VAR_GLOBAL   // PLC tag table "GW_SDC_TO_EMS01_TagTable"
   "SDC_EMS01_Carrier1_Spare0" AT %Q10768.0 : Bool;
   "SDC_EMS01_Carrier1_DriveTripped" AT %Q10768.1 : Bool;
   "SDC_EMS01_Carrier1_Spare2" AT %Q10768.2 : Bool;
   "SDC_EMS01_Carrier1_PositioningComplete" AT %Q10768.3 : Bool;
   "SDC_EMS01_Carrier1_RunStopPressed" AT %Q10768.4 : Bool;
   "SDC_EMS01_Carrier1_Moving" AT %Q10768.5 : Bool;
   "SDC_EMS01_Carrier1_Faulted" AT %Q10768.6 : Bool;
   "SDC_EMS01_Carrier1_InAuto" AT %Q10768.7 : Bool;
   "SDC_EMS01_Carrier2_Spare0" AT %Q10769.0 : Bool;
   "SDC_EMS01_Carrier2_DriveTripped" AT %Q10769.1 : Bool;
   "SDC_EMS01_Carrier2_Spare2" AT %Q10769.2 : Bool;
   "SDC_EMS01_Carrier2_PositioningComplete" AT %Q10769.3 : Bool;
   "SDC_EMS01_Carrier2_RunStopPressed" AT %Q10769.4 : Bool;
   "SDC_EMS01_Carrier2_Moving" AT %Q10769.5 : Bool;
   "SDC_EMS01_Carrier2_Faulted" AT %Q10769.6 : Bool;
   "SDC_EMS01_Carrier2_InAuto" AT %Q10769.7 : Bool;
   "SDC_EMS01_Carrier3_Spare0" AT %Q10770.0 : Bool;
   "SDC_EMS01_Carrier3_DriveTripped" AT %Q10770.1 : Bool;
   "SDC_EMS01_Carrier3_Spare2" AT %Q10770.2 : Bool;
   "SDC_EMS01_Carrier3_PositioningComplete" AT %Q10770.3 : Bool;
   "SDC_EMS01_Carrier3_RunStopPressed" AT %Q10770.4 : Bool;
   "SDC_EMS01_Carrier3_Moving" AT %Q10770.5 : Bool;
   "SDC_EMS01_Carrier3_Faulted" AT %Q10770.6 : Bool;
   "SDC_EMS01_Carrier3_InAuto" AT %Q10770.7 : Bool;
   "SDC_EMS01_Carrier4_Spare0" AT %Q10771.0 : Bool;
   "SDC_EMS01_Carrier4_DriveTripped" AT %Q10771.1 : Bool;
   "SDC_EMS01_Carrier4_Spare2" AT %Q10771.2 : Bool;
   "SDC_EMS01_Carrier4_PositioningComplete" AT %Q10771.3 : Bool;
   "SDC_EMS01_Carrier4_RunStopPressed" AT %Q10771.4 : Bool;
   "SDC_EMS01_Carrier4_Moving" AT %Q10771.5 : Bool;
   "SDC_EMS01_Carrier4_Faulted" AT %Q10771.6 : Bool;
   "SDC_EMS01_Carrier4_InAuto" AT %Q10771.7 : Bool;
   "SDC_EMS01_Carrier5_Spare0" AT %Q10772.0 : Bool;
   "SDC_EMS01_Carrier5_DriveTripped" AT %Q10772.1 : Bool;
   "SDC_EMS01_Carrier5_Spare2" AT %Q10772.2 : Bool;
   "SDC_EMS01_Carrier5_PositioningComplete" AT %Q10772.3 : Bool;
   "SDC_EMS01_Carrier5_RunStopPressed" AT %Q10772.4 : Bool;
   "SDC_EMS01_Carrier5_Moving" AT %Q10772.5 : Bool;
   "SDC_EMS01_Carrier5_Faulted" AT %Q10772.6 : Bool;
   "SDC_EMS01_Carrier5_InAuto" AT %Q10772.7 : Bool;
   "SDC_EMS01_Carrier6_Spare0" AT %Q10773.0 : Bool;
   "SDC_EMS01_Carrier6_DriveTripped" AT %Q10773.1 : Bool;
   "SDC_EMS01_Carrier6_Spare2" AT %Q10773.2 : Bool;
   "SDC_EMS01_Carrier6_PositioningComplete" AT %Q10773.3 : Bool;
   "SDC_EMS01_Carrier6_RunStopPressed" AT %Q10773.4 : Bool;
   "SDC_EMS01_Carrier6_Moving" AT %Q10773.5 : Bool;
   "SDC_EMS01_Carrier6_Faulted" AT %Q10773.6 : Bool;
   "SDC_EMS01_Carrier6_InAuto" AT %Q10773.7 : Bool;
   "SDC_EMS01_Carrier7_Spare0" AT %Q10774.0 : Bool;
   "SDC_EMS01_Carrier7_DriveTripped" AT %Q10774.1 : Bool;
   "SDC_EMS01_Carrier7_Spare2" AT %Q10774.2 : Bool;
   "SDC_EMS01_Carrier7_PositioningComplete" AT %Q10774.3 : Bool;
   "SDC_EMS01_Carrier7_RunStopPressed" AT %Q10774.4 : Bool;
   "SDC_EMS01_Carrier7_Moving" AT %Q10774.5 : Bool;
   "SDC_EMS01_Carrier7_Faulted" AT %Q10774.6 : Bool;
   "SDC_EMS01_Carrier7_InAuto" AT %Q10774.7 : Bool;
   "SDC_EMS01_Carrier8_Spare0" AT %Q10775.0 : Bool;
   "SDC_EMS01_Carrier8_DriveTripped" AT %Q10775.1 : Bool;
   "SDC_EMS01_Carrier8_Spare2" AT %Q10775.2 : Bool;
   "SDC_EMS01_Carrier8_PositioningComplete" AT %Q10775.3 : Bool;
   "SDC_EMS01_Carrier8_RunStopPressed" AT %Q10775.4 : Bool;
   "SDC_EMS01_Carrier8_Moving" AT %Q10775.5 : Bool;
   "SDC_EMS01_Carrier8_Faulted" AT %Q10775.6 : Bool;
   "SDC_EMS01_Carrier8_InAuto" AT %Q10775.7 : Bool;
   "SDC_EMS01_Carrier9_Spare0" AT %Q10776.0 : Bool;
   "SDC_EMS01_Carrier9_DriveTripped" AT %Q10776.1 : Bool;
   "SDC_EMS01_Carrier9_Spare2" AT %Q10776.2 : Bool;
   "SDC_EMS01_Carrier9_PositioningComplete" AT %Q10776.3 : Bool;
   "SDC_EMS01_Carrier9_RunStopPressed" AT %Q10776.4 : Bool;
   "SDC_EMS01_Carrier9_Moving" AT %Q10776.5 : Bool;
   "SDC_EMS01_Carrier9_Faulted" AT %Q10776.6 : Bool;
   "SDC_EMS01_Carrier9_InAuto" AT %Q10776.7 : Bool;
   "SDC_EMS01_Carrier10_Spare0" AT %Q10777.0 : Bool;
   "SDC_EMS01_Carrier10_DriveTripped" AT %Q10777.1 : Bool;
   "SDC_EMS01_Carrier10_Spare2" AT %Q10777.2 : Bool;
   "SDC_EMS01_Carrier10_PositioningComplete" AT %Q10777.3 : Bool;
   "SDC_EMS01_Carrier10_RunStopPressed" AT %Q10777.4 : Bool;
   "SDC_EMS01_Carrier10_Moving" AT %Q10777.5 : Bool;
   "SDC_EMS01_Carrier10_Faulted" AT %Q10777.6 : Bool;
   "SDC_EMS01_Carrier10_InAuto" AT %Q10777.7 : Bool;
   "SDC_EMS01_Carrier11_Spare0" AT %Q10778.0 : Bool;
   "SDC_EMS01_Carrier11_DriveTripped" AT %Q10778.1 : Bool;
   "SDC_EMS01_Carrier11_Spare2" AT %Q10778.2 : Bool;
   "SDC_EMS01_Carrier11_PositioningComplete" AT %Q10778.3 : Bool;
   "SDC_EMS01_Carrier11_RunStopPressed" AT %Q10778.4 : Bool;
   "SDC_EMS01_Carrier11_Moving" AT %Q10778.5 : Bool;
   "SDC_EMS01_Carrier11_Faulted" AT %Q10778.6 : Bool;
   "SDC_EMS01_Carrier11_InAuto" AT %Q10778.7 : Bool;
   "SDC_EMS01_Carrier12_Spare0" AT %Q10779.0 : Bool;
   "SDC_EMS01_Carrier12_DriveTripped" AT %Q10779.1 : Bool;
   "SDC_EMS01_Carrier12_Spare2" AT %Q10779.2 : Bool;
   "SDC_EMS01_Carrier12_PositioningComplete" AT %Q10779.3 : Bool;
   "SDC_EMS01_Carrier12_RunStopPressed" AT %Q10779.4 : Bool;
   "SDC_EMS01_Carrier12_Moving" AT %Q10779.5 : Bool;
   "SDC_EMS01_Carrier12_Faulted" AT %Q10779.6 : Bool;
   "SDC_EMS01_Carrier12_InAuto" AT %Q10779.7 : Bool;
   "SDC_EMS01_Carrier13_Spare0" AT %Q10780.0 : Bool;
   "SDC_EMS01_Carrier13_DriveTripped" AT %Q10780.1 : Bool;
   "SDC_EMS01_Carrier13_Spare2" AT %Q10780.2 : Bool;
   "SDC_EMS01_Carrier13_PositioningComplete" AT %Q10780.3 : Bool;
   "SDC_EMS01_Carrier13_RunStopPressed" AT %Q10780.4 : Bool;
   "SDC_EMS01_Carrier13_Moving" AT %Q10780.5 : Bool;
   "SDC_EMS01_Carrier13_Faulted" AT %Q10780.6 : Bool;
   "SDC_EMS01_Carrier13_InAuto" AT %Q10780.7 : Bool;
   "SDC_EMS01_Carrier14_Spare0" AT %Q10781.0 : Bool;
   "SDC_EMS01_Carrier14_DriveTripped" AT %Q10781.1 : Bool;
   "SDC_EMS01_Carrier14_Spare2" AT %Q10781.2 : Bool;
   "SDC_EMS01_Carrier14_PositioningComplete" AT %Q10781.3 : Bool;
   "SDC_EMS01_Carrier14_RunStopPressed" AT %Q10781.4 : Bool;
   "SDC_EMS01_Carrier14_Moving" AT %Q10781.5 : Bool;
   "SDC_EMS01_Carrier14_Faulted" AT %Q10781.6 : Bool;
   "SDC_EMS01_Carrier14_InAuto" AT %Q10781.7 : Bool;
   "SDC_EMS01_Carrier15_Spare0" AT %Q10782.0 : Bool;
   "SDC_EMS01_Carrier15_DriveTripped" AT %Q10782.1 : Bool;
   "SDC_EMS01_Carrier15_Spare2" AT %Q10782.2 : Bool;
   "SDC_EMS01_Carrier15_PositioningComplete" AT %Q10782.3 : Bool;
   "SDC_EMS01_Carrier15_RunStopPressed" AT %Q10782.4 : Bool;
   "SDC_EMS01_Carrier15_Moving" AT %Q10782.5 : Bool;
   "SDC_EMS01_Carrier15_Faulted" AT %Q10782.6 : Bool;
   "SDC_EMS01_Carrier15_InAuto" AT %Q10782.7 : Bool;
   "SDC_EMS01_Carrier16_Spare0" AT %Q10783.0 : Bool;
   "SDC_EMS01_Carrier16_DriveTripped" AT %Q10783.1 : Bool;
   "SDC_EMS01_Carrier16_Spare2" AT %Q10783.2 : Bool;
   "SDC_EMS01_Carrier16_PositioningComplete" AT %Q10783.3 : Bool;
   "SDC_EMS01_Carrier16_RunStopPressed" AT %Q10783.4 : Bool;
   "SDC_EMS01_Carrier16_Moving" AT %Q10783.5 : Bool;
   "SDC_EMS01_Carrier16_Faulted" AT %Q10783.6 : Bool;
   "SDC_EMS01_Carrier16_InAuto" AT %Q10783.7 : Bool;
   "SDC_EMS01_Carrier17_Spare0" AT %Q10784.0 : Bool;
   "SDC_EMS01_Carrier17_DriveTripped" AT %Q10784.1 : Bool;
   "SDC_EMS01_Carrier17_Spare2" AT %Q10784.2 : Bool;
   "SDC_EMS01_Carrier17_PositioningComplete" AT %Q10784.3 : Bool;
   "SDC_EMS01_Carrier17_RunStopPressed" AT %Q10784.4 : Bool;
   "SDC_EMS01_Carrier17_Moving" AT %Q10784.5 : Bool;
   "SDC_EMS01_Carrier17_Faulted" AT %Q10784.6 : Bool;
   "SDC_EMS01_Carrier17_InAuto" AT %Q10784.7 : Bool;
   "SDC_EMS01_Carrier18_Spare0" AT %Q10785.0 : Bool;
   "SDC_EMS01_Carrier18_DriveTripped" AT %Q10785.1 : Bool;
   "SDC_EMS01_Carrier18_Spare2" AT %Q10785.2 : Bool;
   "SDC_EMS01_Carrier18_PositioningComplete" AT %Q10785.3 : Bool;
   "SDC_EMS01_Carrier18_RunStopPressed" AT %Q10785.4 : Bool;
   "SDC_EMS01_Carrier18_Moving" AT %Q10785.5 : Bool;
   "SDC_EMS01_Carrier18_Faulted" AT %Q10785.6 : Bool;
   "SDC_EMS01_Carrier18_InAuto" AT %Q10785.7 : Bool;
   "SDC_EMS01_Carrier19_Spare0" AT %Q10786.0 : Bool;
   "SDC_EMS01_Carrier19_DriveTripped" AT %Q10786.1 : Bool;
   "SDC_EMS01_Carrier19_Spare2" AT %Q10786.2 : Bool;
   "SDC_EMS01_Carrier19_PositioningComplete" AT %Q10786.3 : Bool;
   "SDC_EMS01_Carrier19_RunStopPressed" AT %Q10786.4 : Bool;
   "SDC_EMS01_Carrier19_Moving" AT %Q10786.5 : Bool;
   "SDC_EMS01_Carrier19_Faulted" AT %Q10786.6 : Bool;
   "SDC_EMS01_Carrier19_InAuto" AT %Q10786.7 : Bool;
   "SDC_EMS01_Carrier20_Spare0" AT %Q10787.0 : Bool;
   "SDC_EMS01_Carrier20_DriveTripped" AT %Q10787.1 : Bool;
   "SDC_EMS01_Carrier20_Spare2" AT %Q10787.2 : Bool;
   "SDC_EMS01_Carrier20_PositioningComplete" AT %Q10787.3 : Bool;
   "SDC_EMS01_Carrier20_RunStopPressed" AT %Q10787.4 : Bool;
   "SDC_EMS01_Carrier20_Moving" AT %Q10787.5 : Bool;
   "SDC_EMS01_Carrier20_Faulted" AT %Q10787.6 : Bool;
   "SDC_EMS01_Carrier20_InAuto" AT %Q10787.7 : Bool;
   "SDC_EMS01_Carrier21_Spare0" AT %Q10788.0 : Bool;
   "SDC_EMS01_Carrier21_DriveTripped" AT %Q10788.1 : Bool;
   "SDC_EMS01_Carrier21_Spare2" AT %Q10788.2 : Bool;
   "SDC_EMS01_Carrier21_PositioningComplete" AT %Q10788.3 : Bool;
   "SDC_EMS01_Carrier21_RunStopPressed" AT %Q10788.4 : Bool;
   "SDC_EMS01_Carrier21_Moving" AT %Q10788.5 : Bool;
   "SDC_EMS01_Carrier21_Faulted" AT %Q10788.6 : Bool;
   "SDC_EMS01_Carrier21_InAuto" AT %Q10788.7 : Bool;
   "SDC_EMS01_Carrier22_Spare0" AT %Q10789.0 : Bool;
   "SDC_EMS01_Carrier22_DriveTripped" AT %Q10789.1 : Bool;
   "SDC_EMS01_Carrier22_Spare2" AT %Q10789.2 : Bool;
   "SDC_EMS01_Carrier22_PositioningComplete" AT %Q10789.3 : Bool;
   "SDC_EMS01_Carrier22_RunStopPressed" AT %Q10789.4 : Bool;
   "SDC_EMS01_Carrier22_Moving" AT %Q10789.5 : Bool;
   "SDC_EMS01_Carrier22_Faulted" AT %Q10789.6 : Bool;
   "SDC_EMS01_Carrier22_InAuto" AT %Q10789.7 : Bool;
   "SDC_EMS01_Carrier23_Spare0" AT %Q10790.0 : Bool;
   "SDC_EMS01_Carrier23_DriveTripped" AT %Q10790.1 : Bool;
   "SDC_EMS01_Carrier23_Spare2" AT %Q10790.2 : Bool;
   "SDC_EMS01_Carrier23_PositioningComplete" AT %Q10790.3 : Bool;
   "SDC_EMS01_Carrier23_RunStopPressed" AT %Q10790.4 : Bool;
   "SDC_EMS01_Carrier23_Moving" AT %Q10790.5 : Bool;
   "SDC_EMS01_Carrier23_Faulted" AT %Q10790.6 : Bool;
   "SDC_EMS01_Carrier23_InAuto" AT %Q10790.7 : Bool;
   "SDC_EMS01_Carrier24_Spare0" AT %Q10791.0 : Bool;
   "SDC_EMS01_Carrier24_DriveTripped" AT %Q10791.1 : Bool;
   "SDC_EMS01_Carrier24_Spare2" AT %Q10791.2 : Bool;
   "SDC_EMS01_Carrier24_PositioningComplete" AT %Q10791.3 : Bool;
   "SDC_EMS01_Carrier24_RunStopPressed" AT %Q10791.4 : Bool;
   "SDC_EMS01_Carrier24_Moving" AT %Q10791.5 : Bool;
   "SDC_EMS01_Carrier24_Faulted" AT %Q10791.6 : Bool;
   "SDC_EMS01_Carrier24_InAuto" AT %Q10791.7 : Bool;
   "SDC_EMS01_Carrier25_Spare0" AT %Q10792.0 : Bool;
   "SDC_EMS01_Carrier25_DriveTripped" AT %Q10792.1 : Bool;
   "SDC_EMS01_Carrier25_Spare2" AT %Q10792.2 : Bool;
   "SDC_EMS01_Carrier25_PositioningComplete" AT %Q10792.3 : Bool;
   "SDC_EMS01_Carrier25_RunStopPressed" AT %Q10792.4 : Bool;
   "SDC_EMS01_Carrier25_Moving" AT %Q10792.5 : Bool;
   "SDC_EMS01_Carrier25_Faulted" AT %Q10792.6 : Bool;
   "SDC_EMS01_Carrier25_InAuto" AT %Q10792.7 : Bool;
   "SDC_EMS01_Carrier26_Spare0" AT %Q10793.0 : Bool;
   "SDC_EMS01_Carrier26_DriveTripped" AT %Q10793.1 : Bool;
   "SDC_EMS01_Carrier26_Spare2" AT %Q10793.2 : Bool;
   "SDC_EMS01_Carrier26_PositioningComplete" AT %Q10793.3 : Bool;
   "SDC_EMS01_Carrier26_RunStopPressed" AT %Q10793.4 : Bool;
   "SDC_EMS01_Carrier26_Moving" AT %Q10793.5 : Bool;
   "SDC_EMS01_Carrier26_Faulted" AT %Q10793.6 : Bool;
   "SDC_EMS01_Carrier26_InAuto" AT %Q10793.7 : Bool;
   "SDC_EMS01_Carrier27_Spare0" AT %Q10794.0 : Bool;
   "SDC_EMS01_Carrier27_DriveTripped" AT %Q10794.1 : Bool;
   "SDC_EMS01_Carrier27_Spare2" AT %Q10794.2 : Bool;
   "SDC_EMS01_Carrier27_PositioningComplete" AT %Q10794.3 : Bool;
   "SDC_EMS01_Carrier27_RunStopPressed" AT %Q10794.4 : Bool;
   "SDC_EMS01_Carrier27_Moving" AT %Q10794.5 : Bool;
   "SDC_EMS01_Carrier27_Faulted" AT %Q10794.6 : Bool;
   "SDC_EMS01_Carrier27_InAuto" AT %Q10794.7 : Bool;
   "SDC_EMS01_Carrier28_Spare0" AT %Q10795.0 : Bool;
   "SDC_EMS01_Carrier28_DriveTripped" AT %Q10795.1 : Bool;
   "SDC_EMS01_Carrier28_Spare2" AT %Q10795.2 : Bool;
   "SDC_EMS01_Carrier28_PositioningComplete" AT %Q10795.3 : Bool;
   "SDC_EMS01_Carrier28_RunStopPressed" AT %Q10795.4 : Bool;
   "SDC_EMS01_Carrier28_Moving" AT %Q10795.5 : Bool;
   "SDC_EMS01_Carrier28_Faulted" AT %Q10795.6 : Bool;
   "SDC_EMS01_Carrier28_InAuto" AT %Q10795.7 : Bool;
   "SDC_EMS01_Carrier29_Spare0" AT %Q10796.0 : Bool;
   "SDC_EMS01_Carrier29_DriveTripped" AT %Q10796.1 : Bool;
   "SDC_EMS01_Carrier29_Spare2" AT %Q10796.2 : Bool;
   "SDC_EMS01_Carrier29_PositioningComplete" AT %Q10796.3 : Bool;
   "SDC_EMS01_Carrier29_RunStopPressed" AT %Q10796.4 : Bool;
   "SDC_EMS01_Carrier29_Moving" AT %Q10796.5 : Bool;
   "SDC_EMS01_Carrier29_Faulted" AT %Q10796.6 : Bool;
   "SDC_EMS01_Carrier29_InAuto" AT %Q10796.7 : Bool;
   "SDC_EMS01_Carrier30_Spare0" AT %Q10797.0 : Bool;
   "SDC_EMS01_Carrier30_DriveTripped" AT %Q10797.1 : Bool;
   "SDC_EMS01_Carrier30_Spare2" AT %Q10797.2 : Bool;
   "SDC_EMS01_Carrier30_PositioningComplete" AT %Q10797.3 : Bool;
   "SDC_EMS01_Carrier30_RunStopPressed" AT %Q10797.4 : Bool;
   "SDC_EMS01_Carrier30_Moving" AT %Q10797.5 : Bool;
   "SDC_EMS01_Carrier30_Faulted" AT %Q10797.6 : Bool;
   "SDC_EMS01_Carrier30_InAuto" AT %Q10797.7 : Bool;
   "SDC_EMS01_Carrier31_Spare0" AT %Q10798.0 : Bool;
   "SDC_EMS01_Carrier31_DriveTripped" AT %Q10798.1 : Bool;
   "SDC_EMS01_Carrier31_Spare2" AT %Q10798.2 : Bool;
   "SDC_EMS01_Carrier31_PositioningComplete" AT %Q10798.3 : Bool;
   "SDC_EMS01_Carrier31_RunStopPressed" AT %Q10798.4 : Bool;
   "SDC_EMS01_Carrier31_Moving" AT %Q10798.5 : Bool;
   "SDC_EMS01_Carrier31_Faulted" AT %Q10798.6 : Bool;
   "SDC_EMS01_Carrier31_InAuto" AT %Q10798.7 : Bool;
   "SDC_EMS01_Carrier32_Spare0" AT %Q10799.0 : Bool;
   "SDC_EMS01_Carrier32_DriveTripped" AT %Q10799.1 : Bool;
   "SDC_EMS01_Carrier32_Spare2" AT %Q10799.2 : Bool;
   "SDC_EMS01_Carrier32_PositioningComplete" AT %Q10799.3 : Bool;
   "SDC_EMS01_Carrier32_RunStopPressed" AT %Q10799.4 : Bool;
   "SDC_EMS01_Carrier32_Moving" AT %Q10799.5 : Bool;
   "SDC_EMS01_Carrier32_Faulted" AT %Q10799.6 : Bool;
   "SDC_EMS01_Carrier32_InAuto" AT %Q10799.7 : Bool;
   "SDC_EMS01_Carrier33_Spare0" AT %Q10800.0 : Bool;
   "SDC_EMS01_Carrier33_DriveTripped" AT %Q10800.1 : Bool;
   "SDC_EMS01_Carrier33_Spare2" AT %Q10800.2 : Bool;
   "SDC_EMS01_Carrier33_PositioningComplete" AT %Q10800.3 : Bool;
   "SDC_EMS01_Carrier33_RunStopPressed" AT %Q10800.4 : Bool;
   "SDC_EMS01_Carrier33_Moving" AT %Q10800.5 : Bool;
   "SDC_EMS01_Carrier33_Faulted" AT %Q10800.6 : Bool;
   "SDC_EMS01_Carrier33_InAuto" AT %Q10800.7 : Bool;
   "SDC_EMS01_Carrier34_Spare0" AT %Q10801.0 : Bool;
   "SDC_EMS01_Carrier34_DriveTripped" AT %Q10801.1 : Bool;
   "SDC_EMS01_Carrier34_Spare2" AT %Q10801.2 : Bool;
   "SDC_EMS01_Carrier34_PositioningComplete" AT %Q10801.3 : Bool;
   "SDC_EMS01_Carrier34_RunStopPressed" AT %Q10801.4 : Bool;
   "SDC_EMS01_Carrier34_Moving" AT %Q10801.5 : Bool;
   "SDC_EMS01_Carrier34_Faulted" AT %Q10801.6 : Bool;
   "SDC_EMS01_Carrier34_InAuto" AT %Q10801.7 : Bool;
   "SDC_EMS01_Carrier35_Spare0" AT %Q10802.0 : Bool;
   "SDC_EMS01_Carrier35_DriveTripped" AT %Q10802.1 : Bool;
   "SDC_EMS01_Carrier35_Spare2" AT %Q10802.2 : Bool;
   "SDC_EMS01_Carrier35_PositioningComplete" AT %Q10802.3 : Bool;
   "SDC_EMS01_Carrier35_RunStopPressed" AT %Q10802.4 : Bool;
   "SDC_EMS01_Carrier35_Moving" AT %Q10802.5 : Bool;
   "SDC_EMS01_Carrier35_Faulted" AT %Q10802.6 : Bool;
   "SDC_EMS01_Carrier35_InAuto" AT %Q10802.7 : Bool;
   "SDC_EMS01_Carrier36_Spare0" AT %Q10803.0 : Bool;
   "SDC_EMS01_Carrier36_DriveTripped" AT %Q10803.1 : Bool;
   "SDC_EMS01_Carrier36_Spare2" AT %Q10803.2 : Bool;
   "SDC_EMS01_Carrier36_PositioningComplete" AT %Q10803.3 : Bool;
   "SDC_EMS01_Carrier36_RunStopPressed" AT %Q10803.4 : Bool;
   "SDC_EMS01_Carrier36_Moving" AT %Q10803.5 : Bool;
   "SDC_EMS01_Carrier36_Faulted" AT %Q10803.6 : Bool;
   "SDC_EMS01_Carrier36_InAuto" AT %Q10803.7 : Bool;
   "SDC_EMS01_Carrier37_Spare0" AT %Q10804.0 : Bool;
   "SDC_EMS01_Carrier37_DriveTripped" AT %Q10804.1 : Bool;
   "SDC_EMS01_Carrier37_Spare2" AT %Q10804.2 : Bool;
   "SDC_EMS01_Carrier37_PositioningComplete" AT %Q10804.3 : Bool;
   "SDC_EMS01_Carrier37_RunStopPressed" AT %Q10804.4 : Bool;
   "SDC_EMS01_Carrier37_Moving" AT %Q10804.5 : Bool;
   "SDC_EMS01_Carrier37_Faulted" AT %Q10804.6 : Bool;
   "SDC_EMS01_Carrier37_InAuto" AT %Q10804.7 : Bool;
   "SDC_EMS01_Carrier38_Spare0" AT %Q10805.0 : Bool;
   "SDC_EMS01_Carrier38_DriveTripped" AT %Q10805.1 : Bool;
   "SDC_EMS01_Carrier38_Spare2" AT %Q10805.2 : Bool;
   "SDC_EMS01_Carrier38_PositioningComplete" AT %Q10805.3 : Bool;
   "SDC_EMS01_Carrier38_RunStopPressed" AT %Q10805.4 : Bool;
   "SDC_EMS01_Carrier38_Moving" AT %Q10805.5 : Bool;
   "SDC_EMS01_Carrier38_Faulted" AT %Q10805.6 : Bool;
   "SDC_EMS01_Carrier38_InAuto" AT %Q10805.7 : Bool;
   "SDC_EMS01_Carrier39_Spare0" AT %Q10806.0 : Bool;
   "SDC_EMS01_Carrier39_DriveTripped" AT %Q10806.1 : Bool;
   "SDC_EMS01_Carrier39_Spare2" AT %Q10806.2 : Bool;
   "SDC_EMS01_Carrier39_PositioningComplete" AT %Q10806.3 : Bool;
   "SDC_EMS01_Carrier39_RunStopPressed" AT %Q10806.4 : Bool;
   "SDC_EMS01_Carrier39_Moving" AT %Q10806.5 : Bool;
   "SDC_EMS01_Carrier39_Faulted" AT %Q10806.6 : Bool;
   "SDC_EMS01_Carrier39_InAuto" AT %Q10806.7 : Bool;
   "SDC_EMS01_Carrier40_Spare0" AT %Q10807.0 : Bool;
   "SDC_EMS01_Carrier40_DriveTripped" AT %Q10807.1 : Bool;
   "SDC_EMS01_Carrier40_Spare2" AT %Q10807.2 : Bool;
   "SDC_EMS01_Carrier40_PositioningComplete" AT %Q10807.3 : Bool;
   "SDC_EMS01_Carrier40_RunStopPressed" AT %Q10807.4 : Bool;
   "SDC_EMS01_Carrier40_Moving" AT %Q10807.5 : Bool;
   "SDC_EMS01_Carrier40_Faulted" AT %Q10807.6 : Bool;
   "SDC_EMS01_Carrier40_InAuto" AT %Q10807.7 : Bool;
   "SDC_EMS01_Carrier41_Spare0" AT %Q10808.0 : Bool;
   "SDC_EMS01_Carrier41_DriveTripped" AT %Q10808.1 : Bool;
   "SDC_EMS01_Carrier41_Spare2" AT %Q10808.2 : Bool;
   "SDC_EMS01_Carrier41_PositioningComplete" AT %Q10808.3 : Bool;
   "SDC_EMS01_Carrier41_RunStopPressed" AT %Q10808.4 : Bool;
   "SDC_EMS01_Carrier41_Moving" AT %Q10808.5 : Bool;
   "SDC_EMS01_Carrier41_Faulted" AT %Q10808.6 : Bool;
   "SDC_EMS01_Carrier41_InAuto" AT %Q10808.7 : Bool;
   "SDC_EMS01_Carrier42_Spare0" AT %Q10809.0 : Bool;
   "SDC_EMS01_Carrier42_DriveTripped" AT %Q10809.1 : Bool;
   "SDC_EMS01_Carrier42_Spare2" AT %Q10809.2 : Bool;
   "SDC_EMS01_Carrier42_PositioningComplete" AT %Q10809.3 : Bool;
   "SDC_EMS01_Carrier42_RunStopPressed" AT %Q10809.4 : Bool;
   "SDC_EMS01_Carrier42_Moving" AT %Q10809.5 : Bool;
   "SDC_EMS01_Carrier42_Faulted" AT %Q10809.6 : Bool;
   "SDC_EMS01_Carrier42_InAuto" AT %Q10809.7 : Bool;
   "SDC_EMS01_Carrier43_Spare0" AT %Q10810.0 : Bool;
   "SDC_EMS01_Carrier43_DriveTripped" AT %Q10810.1 : Bool;
   "SDC_EMS01_Carrier43_Spare2" AT %Q10810.2 : Bool;
   "SDC_EMS01_Carrier43_PositioningComplete" AT %Q10810.3 : Bool;
   "SDC_EMS01_Carrier43_RunStopPressed" AT %Q10810.4 : Bool;
   "SDC_EMS01_Carrier43_Moving" AT %Q10810.5 : Bool;
   "SDC_EMS01_Carrier43_Faulted" AT %Q10810.6 : Bool;
   "SDC_EMS01_Carrier43_InAuto" AT %Q10810.7 : Bool;
   "SDC_EMS01_Carrier44_Spare0" AT %Q10811.0 : Bool;
   "SDC_EMS01_Carrier44_DriveTripped" AT %Q10811.1 : Bool;
   "SDC_EMS01_Carrier44_Spare2" AT %Q10811.2 : Bool;
   "SDC_EMS01_Carrier44_PositioningComplete" AT %Q10811.3 : Bool;
   "SDC_EMS01_Carrier44_RunStopPressed" AT %Q10811.4 : Bool;
   "SDC_EMS01_Carrier44_Moving" AT %Q10811.5 : Bool;
   "SDC_EMS01_Carrier44_Faulted" AT %Q10811.6 : Bool;
   "SDC_EMS01_Carrier44_InAuto" AT %Q10811.7 : Bool;
   "SDC_EMS01_Carrier45_Spare0" AT %Q10812.0 : Bool;
   "SDC_EMS01_Carrier45_DriveTripped" AT %Q10812.1 : Bool;
   "SDC_EMS01_Carrier45_Spare2" AT %Q10812.2 : Bool;
   "SDC_EMS01_Carrier45_PositioningComplete" AT %Q10812.3 : Bool;
   "SDC_EMS01_Carrier45_RunStopPressed" AT %Q10812.4 : Bool;
   "SDC_EMS01_Carrier45_Moving" AT %Q10812.5 : Bool;
   "SDC_EMS01_Carrier45_Faulted" AT %Q10812.6 : Bool;
   "SDC_EMS01_Carrier45_InAuto" AT %Q10812.7 : Bool;
   "SDC_EMS01_Carrier46_Spare0" AT %Q10813.0 : Bool;
   "SDC_EMS01_Carrier46_DriveTripped" AT %Q10813.1 : Bool;
   "SDC_EMS01_Carrier46_Spare2" AT %Q10813.2 : Bool;
   "SDC_EMS01_Carrier46_PositioningComplete" AT %Q10813.3 : Bool;
   "SDC_EMS01_Carrier46_RunStopPressed" AT %Q10813.4 : Bool;
   "SDC_EMS01_Carrier46_Moving" AT %Q10813.5 : Bool;
   "SDC_EMS01_Carrier46_Faulted" AT %Q10813.6 : Bool;
   "SDC_EMS01_Carrier46_InAuto" AT %Q10813.7 : Bool;
   "SDC_EMS01_Carrier47_Spare0" AT %Q10814.0 : Bool;
   "SDC_EMS01_Carrier47_DriveTripped" AT %Q10814.1 : Bool;
   "SDC_EMS01_Carrier47_Spare2" AT %Q10814.2 : Bool;
   "SDC_EMS01_Carrier47_PositioningComplete" AT %Q10814.3 : Bool;
   "SDC_EMS01_Carrier47_RunStopPressed" AT %Q10814.4 : Bool;
   "SDC_EMS01_Carrier47_Moving" AT %Q10814.5 : Bool;
   "SDC_EMS01_Carrier47_Faulted" AT %Q10814.6 : Bool;
   "SDC_EMS01_Carrier47_InAuto" AT %Q10814.7 : Bool;
   "SDC_EMS01_Carrier48_Spare0" AT %Q10815.0 : Bool;
   "SDC_EMS01_Carrier48_DriveTripped" AT %Q10815.1 : Bool;
   "SDC_EMS01_Carrier48_Spare2" AT %Q10815.2 : Bool;
   "SDC_EMS01_Carrier48_PositioningComplete" AT %Q10815.3 : Bool;
   "SDC_EMS01_Carrier48_RunStopPressed" AT %Q10815.4 : Bool;
   "SDC_EMS01_Carrier48_Moving" AT %Q10815.5 : Bool;
   "SDC_EMS01_Carrier48_Faulted" AT %Q10815.6 : Bool;
   "SDC_EMS01_Carrier48_InAuto" AT %Q10815.7 : Bool;
   "SDC_EMS01_Carrier49_Spare0" AT %Q10816.0 : Bool;
   "SDC_EMS01_Carrier49_DriveTripped" AT %Q10816.1 : Bool;
   "SDC_EMS01_Carrier49_Spare2" AT %Q10816.2 : Bool;
   "SDC_EMS01_Carrier49_PositioningComplete" AT %Q10816.3 : Bool;
   "SDC_EMS01_Carrier49_RunStopPressed" AT %Q10816.4 : Bool;
   "SDC_EMS01_Carrier49_Moving" AT %Q10816.5 : Bool;
   "SDC_EMS01_Carrier49_Faulted" AT %Q10816.6 : Bool;
   "SDC_EMS01_Carrier49_InAuto" AT %Q10816.7 : Bool;
   "SDC_EMS01_Carrier50_Spare0" AT %Q10817.0 : Bool;
   "SDC_EMS01_Carrier50_DriveTripped" AT %Q10817.1 : Bool;
   "SDC_EMS01_Carrier50_Spare2" AT %Q10817.2 : Bool;
   "SDC_EMS01_Carrier50_PositioningComplete" AT %Q10817.3 : Bool;
   "SDC_EMS01_Carrier50_RunStopPressed" AT %Q10817.4 : Bool;
   "SDC_EMS01_Carrier50_Moving" AT %Q10817.5 : Bool;
   "SDC_EMS01_Carrier50_Faulted" AT %Q10817.6 : Bool;
   "SDC_EMS01_Carrier50_InAuto" AT %Q10817.7 : Bool;
   "SDC_EMS01_Carrier51_Spare0" AT %Q10818.0 : Bool;
   "SDC_EMS01_Carrier51_DriveTripped" AT %Q10818.1 : Bool;
   "SDC_EMS01_Carrier51_Spare2" AT %Q10818.2 : Bool;
   "SDC_EMS01_Carrier51_PositioningComplete" AT %Q10818.3 : Bool;
   "SDC_EMS01_Carrier51_RunStopPressed" AT %Q10818.4 : Bool;
   "SDC_EMS01_Carrier51_Moving" AT %Q10818.5 : Bool;
   "SDC_EMS01_Carrier51_Faulted" AT %Q10818.6 : Bool;
   "SDC_EMS01_Carrier51_InAuto" AT %Q10818.7 : Bool;
   "SDC_EMS01_Carrier52_Spare0" AT %Q10819.0 : Bool;
   "SDC_EMS01_Carrier52_DriveTripped" AT %Q10819.1 : Bool;
   "SDC_EMS01_Carrier52_Spare2" AT %Q10819.2 : Bool;
   "SDC_EMS01_Carrier52_PositioningComplete" AT %Q10819.3 : Bool;
   "SDC_EMS01_Carrier52_RunStopPressed" AT %Q10819.4 : Bool;
   "SDC_EMS01_Carrier52_Moving" AT %Q10819.5 : Bool;
   "SDC_EMS01_Carrier52_Faulted" AT %Q10819.6 : Bool;
   "SDC_EMS01_Carrier52_InAuto" AT %Q10819.7 : Bool;
   "SDC_EMS01_Carrier53_Spare0" AT %Q10820.0 : Bool;
   "SDC_EMS01_Carrier53_DriveTripped" AT %Q10820.1 : Bool;
   "SDC_EMS01_Carrier53_Spare2" AT %Q10820.2 : Bool;
   "SDC_EMS01_Carrier53_PositioningComplete" AT %Q10820.3 : Bool;
   "SDC_EMS01_Carrier53_RunStopPressed" AT %Q10820.4 : Bool;
   "SDC_EMS01_Carrier53_Moving" AT %Q10820.5 : Bool;
   "SDC_EMS01_Carrier53_Faulted" AT %Q10820.6 : Bool;
   "SDC_EMS01_Carrier53_InAuto" AT %Q10820.7 : Bool;
   "SDC_EMS01_Carrier54_Spare0" AT %Q10821.0 : Bool;
   "SDC_EMS01_Carrier54_DriveTripped" AT %Q10821.1 : Bool;
   "SDC_EMS01_Carrier54_Spare2" AT %Q10821.2 : Bool;
   "SDC_EMS01_Carrier54_PositioningComplete" AT %Q10821.3 : Bool;
   "SDC_EMS01_Carrier54_RunStopPressed" AT %Q10821.4 : Bool;
   "SDC_EMS01_Carrier54_Moving" AT %Q10821.5 : Bool;
   "SDC_EMS01_Carrier54_Faulted" AT %Q10821.6 : Bool;
   "SDC_EMS01_Carrier54_InAuto" AT %Q10821.7 : Bool;
   "SDC_EMS01_Carrier55_Spare0" AT %Q10822.0 : Bool;
   "SDC_EMS01_Carrier55_DriveTripped" AT %Q10822.1 : Bool;
   "SDC_EMS01_Carrier55_Spare2" AT %Q10822.2 : Bool;
   "SDC_EMS01_Carrier55_PositioningComplete" AT %Q10822.3 : Bool;
   "SDC_EMS01_Carrier55_RunStopPressed" AT %Q10822.4 : Bool;
   "SDC_EMS01_Carrier55_Moving" AT %Q10822.5 : Bool;
   "SDC_EMS01_Carrier55_Faulted" AT %Q10822.6 : Bool;
   "SDC_EMS01_Carrier55_InAuto" AT %Q10822.7 : Bool;
   "SDC_EMS01_Carrier56_Spare0" AT %Q10823.0 : Bool;
   "SDC_EMS01_Carrier56_DriveTripped" AT %Q10823.1 : Bool;
   "SDC_EMS01_Carrier56_Spare2" AT %Q10823.2 : Bool;
   "SDC_EMS01_Carrier56_PositioningComplete" AT %Q10823.3 : Bool;
   "SDC_EMS01_Carrier56_RunStopPressed" AT %Q10823.4 : Bool;
   "SDC_EMS01_Carrier56_Moving" AT %Q10823.5 : Bool;
   "SDC_EMS01_Carrier56_Faulted" AT %Q10823.6 : Bool;
   "SDC_EMS01_Carrier56_InAuto" AT %Q10823.7 : Bool;
   "SDC_EMS01_Carrier57_Spare0" AT %Q10824.0 : Bool;
   "SDC_EMS01_Carrier57_DriveTripped" AT %Q10824.1 : Bool;
   "SDC_EMS01_Carrier57_Spare2" AT %Q10824.2 : Bool;
   "SDC_EMS01_Carrier57_PositioningComplete" AT %Q10824.3 : Bool;
   "SDC_EMS01_Carrier57_RunStopPressed" AT %Q10824.4 : Bool;
   "SDC_EMS01_Carrier57_Moving" AT %Q10824.5 : Bool;
   "SDC_EMS01_Carrier57_Faulted" AT %Q10824.6 : Bool;
   "SDC_EMS01_Carrier57_InAuto" AT %Q10824.7 : Bool;
   "SDC_EMS01_Carrier58_Spare0" AT %Q10825.0 : Bool;
   "SDC_EMS01_Carrier58_DriveTripped" AT %Q10825.1 : Bool;
   "SDC_EMS01_Carrier58_Spare2" AT %Q10825.2 : Bool;
   "SDC_EMS01_Carrier58_PositioningComplete" AT %Q10825.3 : Bool;
   "SDC_EMS01_Carrier58_RunStopPressed" AT %Q10825.4 : Bool;
   "SDC_EMS01_Carrier58_Moving" AT %Q10825.5 : Bool;
   "SDC_EMS01_Carrier58_Faulted" AT %Q10825.6 : Bool;
   "SDC_EMS01_Carrier58_InAuto" AT %Q10825.7 : Bool;
   "SDC_EMS01_Carrier59_Spare0" AT %Q10826.0 : Bool;
   "SDC_EMS01_Carrier59_DriveTripped" AT %Q10826.1 : Bool;
   "SDC_EMS01_Carrier59_Spare2" AT %Q10826.2 : Bool;
   "SDC_EMS01_Carrier59_PositioningComplete" AT %Q10826.3 : Bool;
   "SDC_EMS01_Carrier59_RunStopPressed" AT %Q10826.4 : Bool;
   "SDC_EMS01_Carrier59_Moving" AT %Q10826.5 : Bool;
   "SDC_EMS01_Carrier59_Faulted" AT %Q10826.6 : Bool;
   "SDC_EMS01_Carrier59_InAuto" AT %Q10826.7 : Bool;
   "SDC_EMS01_Carrier60_Spare0" AT %Q10827.0 : Bool;
   "SDC_EMS01_Carrier60_DriveTripped" AT %Q10827.1 : Bool;
   "SDC_EMS01_Carrier60_Spare2" AT %Q10827.2 : Bool;
   "SDC_EMS01_Carrier60_PositioningComplete" AT %Q10827.3 : Bool;
   "SDC_EMS01_Carrier60_RunStopPressed" AT %Q10827.4 : Bool;
   "SDC_EMS01_Carrier60_Moving" AT %Q10827.5 : Bool;
   "SDC_EMS01_Carrier60_Faulted" AT %Q10827.6 : Bool;
   "SDC_EMS01_Carrier60_InAuto" AT %Q10827.7 : Bool;
   "SDC_EMS01_Carrier61_Spare0" AT %Q10828.0 : Bool;
   "SDC_EMS01_Carrier61_DriveTripped" AT %Q10828.1 : Bool;
   "SDC_EMS01_Carrier61_Spare2" AT %Q10828.2 : Bool;
   "SDC_EMS01_Carrier61_PositioningComplete" AT %Q10828.3 : Bool;
   "SDC_EMS01_Carrier61_RunStopPressed" AT %Q10828.4 : Bool;
   "SDC_EMS01_Carrier61_Moving" AT %Q10828.5 : Bool;
   "SDC_EMS01_Carrier61_Faulted" AT %Q10828.6 : Bool;
   "SDC_EMS01_Carrier61_InAuto" AT %Q10828.7 : Bool;
   "SDC_EMS01_Carrier62_Spare0" AT %Q10829.0 : Bool;
   "SDC_EMS01_Carrier62_DriveTripped" AT %Q10829.1 : Bool;
   "SDC_EMS01_Carrier62_Spare2" AT %Q10829.2 : Bool;
   "SDC_EMS01_Carrier62_PositioningComplete" AT %Q10829.3 : Bool;
   "SDC_EMS01_Carrier62_RunStopPressed" AT %Q10829.4 : Bool;
   "SDC_EMS01_Carrier62_Moving" AT %Q10829.5 : Bool;
   "SDC_EMS01_Carrier62_Faulted" AT %Q10829.6 : Bool;
   "SDC_EMS01_Carrier62_InAuto" AT %Q10829.7 : Bool;
   "SDC_EMS01_Carrier63_Spare0" AT %Q10830.0 : Bool;
   "SDC_EMS01_Carrier63_DriveTripped" AT %Q10830.1 : Bool;
   "SDC_EMS01_Carrier63_Spare2" AT %Q10830.2 : Bool;
   "SDC_EMS01_Carrier63_PositioningComplete" AT %Q10830.3 : Bool;
   "SDC_EMS01_Carrier63_RunStopPressed" AT %Q10830.4 : Bool;
   "SDC_EMS01_Carrier63_Moving" AT %Q10830.5 : Bool;
   "SDC_EMS01_Carrier63_Faulted" AT %Q10830.6 : Bool;
   "SDC_EMS01_Carrier63_InAuto" AT %Q10830.7 : Bool;
   "SDC_EMS01_Carrier64_Spare0" AT %Q10831.0 : Bool;
   "SDC_EMS01_Carrier64_DriveTripped" AT %Q10831.1 : Bool;
   "SDC_EMS01_Carrier64_Spare2" AT %Q10831.2 : Bool;
   "SDC_EMS01_Carrier64_PositioningComplete" AT %Q10831.3 : Bool;
   "SDC_EMS01_Carrier64_RunStopPressed" AT %Q10831.4 : Bool;
   "SDC_EMS01_Carrier64_Moving" AT %Q10831.5 : Bool;
   "SDC_EMS01_Carrier64_Faulted" AT %Q10831.6 : Bool;
   "SDC_EMS01_Carrier64_InAuto" AT %Q10831.7 : Bool;
   "SDC_EMS01_Carrier65_Spare0" AT %Q10832.0 : Bool;
   "SDC_EMS01_Carrier65_DriveTripped" AT %Q10832.1 : Bool;
   "SDC_EMS01_Carrier65_Spare2" AT %Q10832.2 : Bool;
   "SDC_EMS01_Carrier65_PositioningComplete" AT %Q10832.3 : Bool;
   "SDC_EMS01_Carrier65_RunStopPressed" AT %Q10832.4 : Bool;
   "SDC_EMS01_Carrier65_Moving" AT %Q10832.5 : Bool;
   "SDC_EMS01_Carrier65_Faulted" AT %Q10832.6 : Bool;
   "SDC_EMS01_Carrier65_InAuto" AT %Q10832.7 : Bool;
   "SDC_EMS01_Carrier66_Spare0" AT %Q10833.0 : Bool;
   "SDC_EMS01_Carrier66_DriveTripped" AT %Q10833.1 : Bool;
   "SDC_EMS01_Carrier66_Spare2" AT %Q10833.2 : Bool;
   "SDC_EMS01_Carrier66_PositioningComplete" AT %Q10833.3 : Bool;
   "SDC_EMS01_Carrier66_RunStopPressed" AT %Q10833.4 : Bool;
   "SDC_EMS01_Carrier66_Moving" AT %Q10833.5 : Bool;
   "SDC_EMS01_Carrier66_Faulted" AT %Q10833.6 : Bool;
   "SDC_EMS01_Carrier66_InAuto" AT %Q10833.7 : Bool;
   "SDC_EMS01_Carrier67_Spare0" AT %Q10834.0 : Bool;
   "SDC_EMS01_Carrier67_DriveTripped" AT %Q10834.1 : Bool;
   "SDC_EMS01_Carrier67_Spare2" AT %Q10834.2 : Bool;
   "SDC_EMS01_Carrier67_PositioningComplete" AT %Q10834.3 : Bool;
   "SDC_EMS01_Carrier67_RunStopPressed" AT %Q10834.4 : Bool;
   "SDC_EMS01_Carrier67_Moving" AT %Q10834.5 : Bool;
   "SDC_EMS01_Carrier67_Faulted" AT %Q10834.6 : Bool;
   "SDC_EMS01_Carrier67_InAuto" AT %Q10834.7 : Bool;
   "SDC_EMS01_Carrier68_Spare0" AT %Q10835.0 : Bool;
   "SDC_EMS01_Carrier68_DriveTripped" AT %Q10835.1 : Bool;
   "SDC_EMS01_Carrier68_Spare2" AT %Q10835.2 : Bool;
   "SDC_EMS01_Carrier68_PositioningComplete" AT %Q10835.3 : Bool;
   "SDC_EMS01_Carrier68_RunStopPressed" AT %Q10835.4 : Bool;
   "SDC_EMS01_Carrier68_Moving" AT %Q10835.5 : Bool;
   "SDC_EMS01_Carrier68_Faulted" AT %Q10835.6 : Bool;
   "SDC_EMS01_Carrier68_InAuto" AT %Q10835.7 : Bool;
   "SDC_EMS01_Carrier69_Spare0" AT %Q10836.0 : Bool;
   "SDC_EMS01_Carrier69_DriveTripped" AT %Q10836.1 : Bool;
   "SDC_EMS01_Carrier69_Spare2" AT %Q10836.2 : Bool;
   "SDC_EMS01_Carrier69_PositioningComplete" AT %Q10836.3 : Bool;
   "SDC_EMS01_Carrier69_RunStopPressed" AT %Q10836.4 : Bool;
   "SDC_EMS01_Carrier69_Moving" AT %Q10836.5 : Bool;
   "SDC_EMS01_Carrier69_Faulted" AT %Q10836.6 : Bool;
   "SDC_EMS01_Carrier69_InAuto" AT %Q10836.7 : Bool;
   "SDC_EMS01_Carrier70_Spare0" AT %Q10837.0 : Bool;
   "SDC_EMS01_Carrier70_DriveTripped" AT %Q10837.1 : Bool;
   "SDC_EMS01_Carrier70_Spare2" AT %Q10837.2 : Bool;
   "SDC_EMS01_Carrier70_PositioningComplete" AT %Q10837.3 : Bool;
   "SDC_EMS01_Carrier70_RunStopPressed" AT %Q10837.4 : Bool;
   "SDC_EMS01_Carrier70_Moving" AT %Q10837.5 : Bool;
   "SDC_EMS01_Carrier70_Faulted" AT %Q10837.6 : Bool;
   "SDC_EMS01_Carrier70_InAuto" AT %Q10837.7 : Bool;
   "SDC_EMS01_Carrier71_Spare0" AT %Q10838.0 : Bool;
   "SDC_EMS01_Carrier71_DriveTripped" AT %Q10838.1 : Bool;
   "SDC_EMS01_Carrier71_Spare2" AT %Q10838.2 : Bool;
   "SDC_EMS01_Carrier71_PositioningComplete" AT %Q10838.3 : Bool;
   "SDC_EMS01_Carrier71_RunStopPressed" AT %Q10838.4 : Bool;
   "SDC_EMS01_Carrier71_Moving" AT %Q10838.5 : Bool;
   "SDC_EMS01_Carrier71_Faulted" AT %Q10838.6 : Bool;
   "SDC_EMS01_Carrier71_InAuto" AT %Q10838.7 : Bool;
   "SDC_EMS01_Carrier72_Spare0" AT %Q10839.0 : Bool;
   "SDC_EMS01_Carrier72_DriveTripped" AT %Q10839.1 : Bool;
   "SDC_EMS01_Carrier72_Spare2" AT %Q10839.2 : Bool;
   "SDC_EMS01_Carrier72_PositioningComplete" AT %Q10839.3 : Bool;
   "SDC_EMS01_Carrier72_RunStopPressed" AT %Q10839.4 : Bool;
   "SDC_EMS01_Carrier72_Moving" AT %Q10839.5 : Bool;
   "SDC_EMS01_Carrier72_Faulted" AT %Q10839.6 : Bool;
   "SDC_EMS01_Carrier72_InAuto" AT %Q10839.7 : Bool;
   "SDC_EMS01_Carrier73_Spare0" AT %Q10840.0 : Bool;
   "SDC_EMS01_Carrier73_DriveTripped" AT %Q10840.1 : Bool;
   "SDC_EMS01_Carrier73_Spare2" AT %Q10840.2 : Bool;
   "SDC_EMS01_Carrier73_PositioningComplete" AT %Q10840.3 : Bool;
   "SDC_EMS01_Carrier73_RunStopPressed" AT %Q10840.4 : Bool;
   "SDC_EMS01_Carrier73_Moving" AT %Q10840.5 : Bool;
   "SDC_EMS01_Carrier73_Faulted" AT %Q10840.6 : Bool;
   "SDC_EMS01_Carrier73_InAuto" AT %Q10840.7 : Bool;
   "SDC_EMS01_Carrier74_Spare0" AT %Q10841.0 : Bool;
   "SDC_EMS01_Carrier74_DriveTripped" AT %Q10841.1 : Bool;
   "SDC_EMS01_Carrier74_Spare2" AT %Q10841.2 : Bool;
   "SDC_EMS01_Carrier74_PositioningComplete" AT %Q10841.3 : Bool;
   "SDC_EMS01_Carrier74_RunStopPressed" AT %Q10841.4 : Bool;
   "SDC_EMS01_Carrier74_Moving" AT %Q10841.5 : Bool;